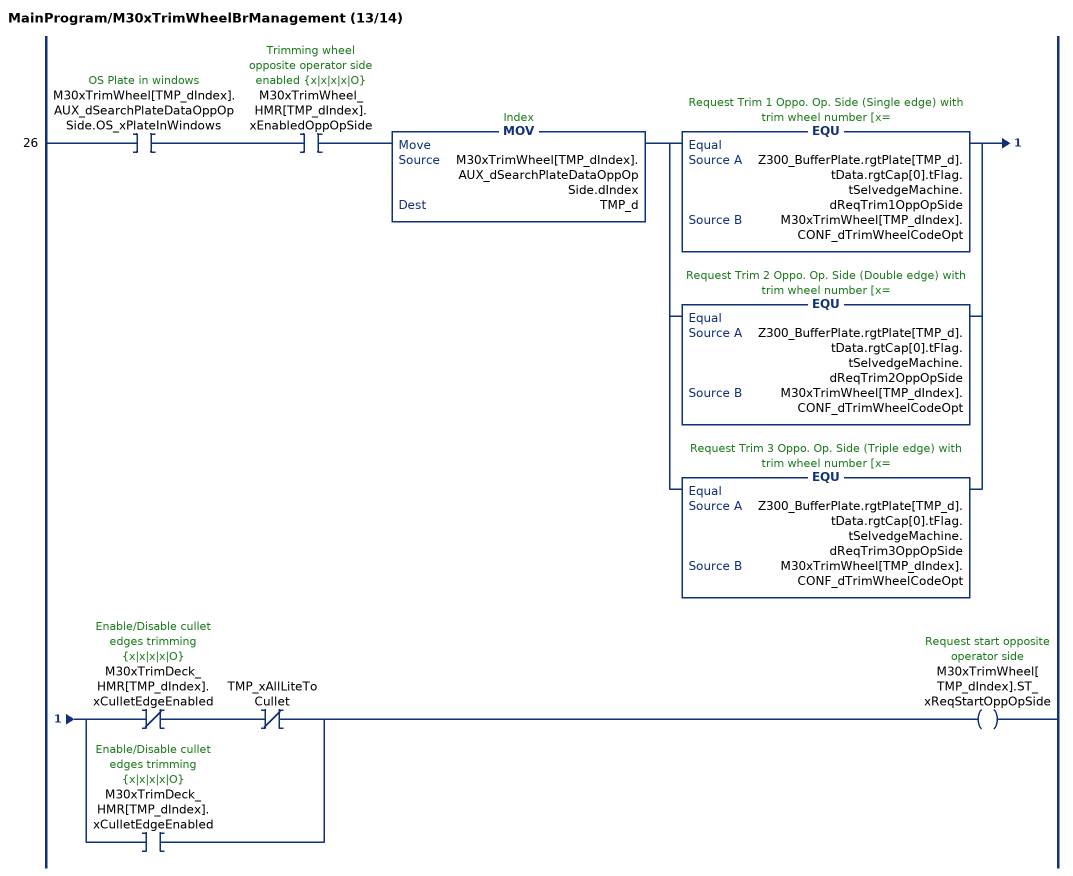
   26: XIC(M30xTrimWheel[TMP_dIndex].AUX_dSearchPlateDataOppOpSide.OS_xPlateInWindows)XIC(M30xTrimWheel_HMR[TMP_dIndex].xEnabledOppOpSide)MOV(M30xTrimWheel[TMP_dIndex].AUX_dSearchPlateDataOppOpSide.dIndex,TMP_d)[EQU(Z300_BufferPlate.rgtPlate[TMP_d].tData.rgtCap[0].tFlag.tSelvedgeMachine.dReqTrim1OppOpSide,M30xTrimWheel[TMP_dIndex].CONF_dTrimWheelCodeOpt) ,EQU(Z300_BufferPlate.rgtPlate[TMP_d].tData.rgtCap[0].tFlag.tSelvedgeMachine.dReqTrim2OppOpSide,M30xTrimWheel[TMP_dIndex].CONF_dTrimWheelCodeOpt) ,EQU(Z300_BufferPlate.rgtPlate[TMP_d].tData.rgtCap[0].tFlag.tSelvedgeMachine.dReqTrim3OppOpSide,M30xTrimWheel[TMP_dIndex].CONF_dTrimWheelCodeOpt) ][XIO(M30xTrimDeck_HMR[TMP_dIndex].xCulletEdgeEnabled) XIO(TMP_xAllLiteToCullet) ,XIC(M30xTrimDeck_HMR[TMP_dIndex].xCulletEdgeEnabled) ]OTE(M30xTrimWheel[TMP_dIndex].ST_xReqStartOppOpSide);
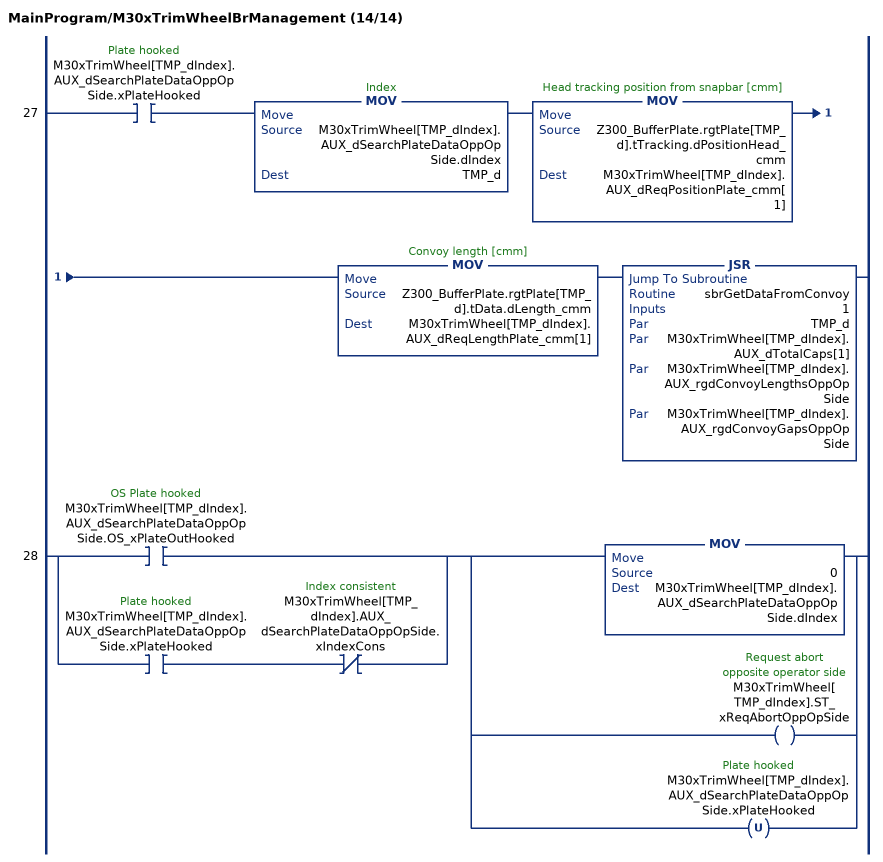
   27: XIC(M30xTrimWheel[TMP_dIndex].AUX_dSearchPlateDataOppOpSide.xPlateHooked)MOV(M30xTrimWheel[TMP_dIndex].AUX_dSearchPlateDataOppOpSide.dIndex,TMP_d)MOV(Z300_BufferPlate.rgtPlate[TMP_d].tTracking.dPositionHead_cmm,M30xTrimWheel[TMP_dIndex].AUX_dReqPositionPlate_cmm[1])MOV(Z300_BufferPlate.rgtPlate[TMP_d].tData.dLength_cmm,M30xTrimWheel[TMP_dIndex].AUX_dReqLengthPlate_cmm[1])JSR(sbrGetDataFromConvoy,1,TMP_d,M30xTrimWheel[TMP_dIndex].AUX_dTotalCaps[1],M30xTrimWheel[TMP_dIndex].AUX_rgdConvoyLengthsOppOpSide,M30xTrimWheel[TMP_dIndex].AUX_rgdConvoyGapsOppOpSide);
   28: [XIC(M30xTrimWheel[TMP_dIndex].AUX_dSearchPlateDataOppOpSide.OS_xPlateOutHooked) ,XIC(M30xTrimWheel[TMP_dIndex].AUX_dSearchPlateDataOppOpSide.xPlateHooked) XIO(M30xTrimWheel[TMP_dIndex].AUX_dSearchPlateDataOppOpSide.xIndexCons) ][MOV(0,M30xTrimWheel[TMP_dIndex].AUX_dSearchPlateDataOppOpSide.dIndex) ,OTE(M30xTrimWheel[TMP_dIndex].ST_xReqAbortOppOpSide) ,OTU(M30xTrimWheel[TMP_dIndex].AUX_dSearchPlateDataOppOpSide.xPlateHooked) ];
END_ROUTINE

ROUTINE M30xTrimWheelTrManagement   (* ladder *)
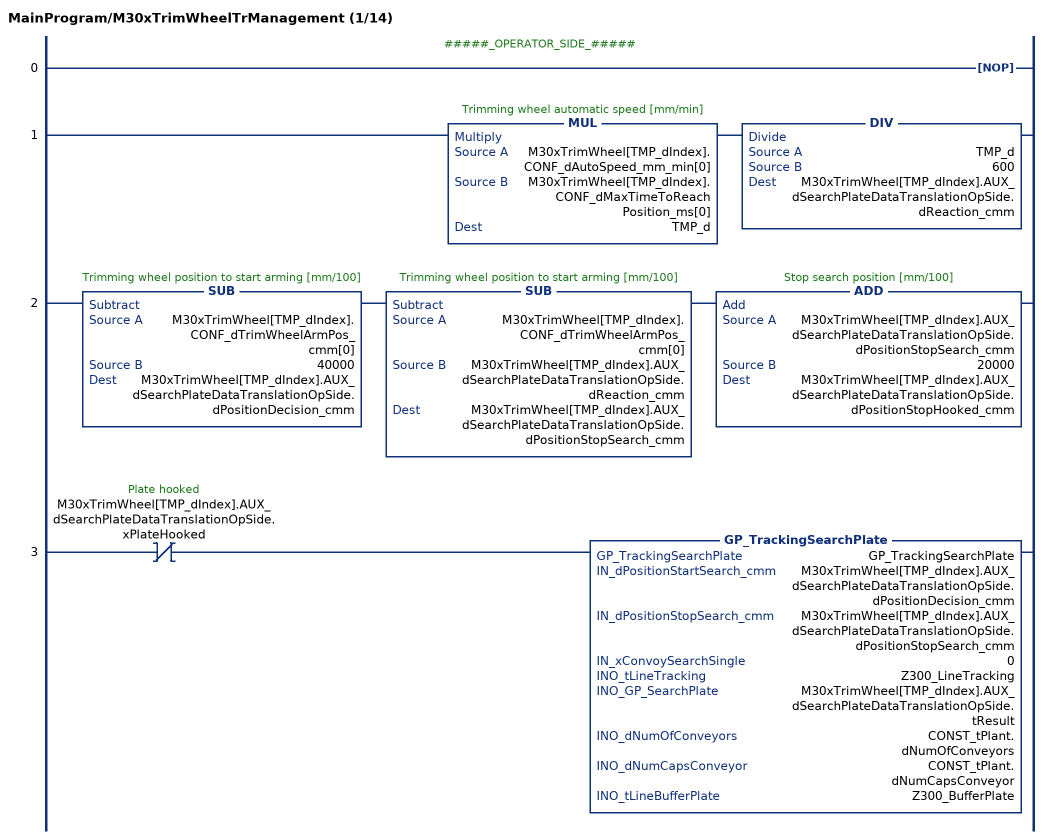
   // #####_OPERATOR_SIDE_#####
   0: NOP();
   1: MUL(M30xTrimWheel[TMP_dIndex].CONF_dAutoSpeed_mm_min[0],M30xTrimWheel[TMP_dIndex].CONF_dMaxTimeToReachPosition_ms[0],TMP_d)DIV(TMP_d,600,M30xTrimWheel[TMP_dIndex].AUX_dSearchPlateDataTranslationOpSide.dReaction_cmm);
   2: SUB(M30xTrimWheel[TMP_dIndex].CONF_dTrimWheelArmPos_cmm[0],40000,M30xTrimWheel[TMP_dIndex].AUX_dSearchPlateDataTranslationOpSide.dPositionDecision_cmm)SUB(M30xTrimWheel[TMP_dIndex].CONF_dTrimWheelArmPos_cmm[0],M30xTrimWheel[TMP_dIndex].AUX_dSearchPlateDataTranslationOpSide.dReaction_cmm,M30xTrimWheel[TMP_dIndex].AUX_dSearchPlateDataTranslationOpSide.dPositionStopSearch_cmm)ADD(M30xTrimWheel[TMP_dIndex].AUX_dSearchPlateDataTranslationOpSide.dPositionStopSearch_cmm,20000,M30xTrimWheel[TMP_dIndex].AUX_dSearchPlateDataTranslationOpSide.dPositionStopHooked_cmm);
   3: XIO(M30xTrimWheel[TMP_dIndex].AUX_dSearchPlateDataTranslationOpSide.xPlateHooked)GP_TrackingSearchPlate(GP_TrackingSearchPlate,M30xTrimWheel[TMP_dIndex].AUX_dSearchPlateDataTranslationOpSide.dPositionDecision_cmm,M30xTrimWheel[TMP_dIndex].AUX_dSearchPlateDataTranslationOpSide.dPositionStopSearch_cmm,0,Z300_LineTracking,M30xTrimWheel[TMP_dIndex].AUX_dSearchPlateDataTranslationOpSide.tResult,CONST_tPlant.dNumOfConveyors,CONST_tPlant.dNumCapsConveyor,Z300_BufferPlate);
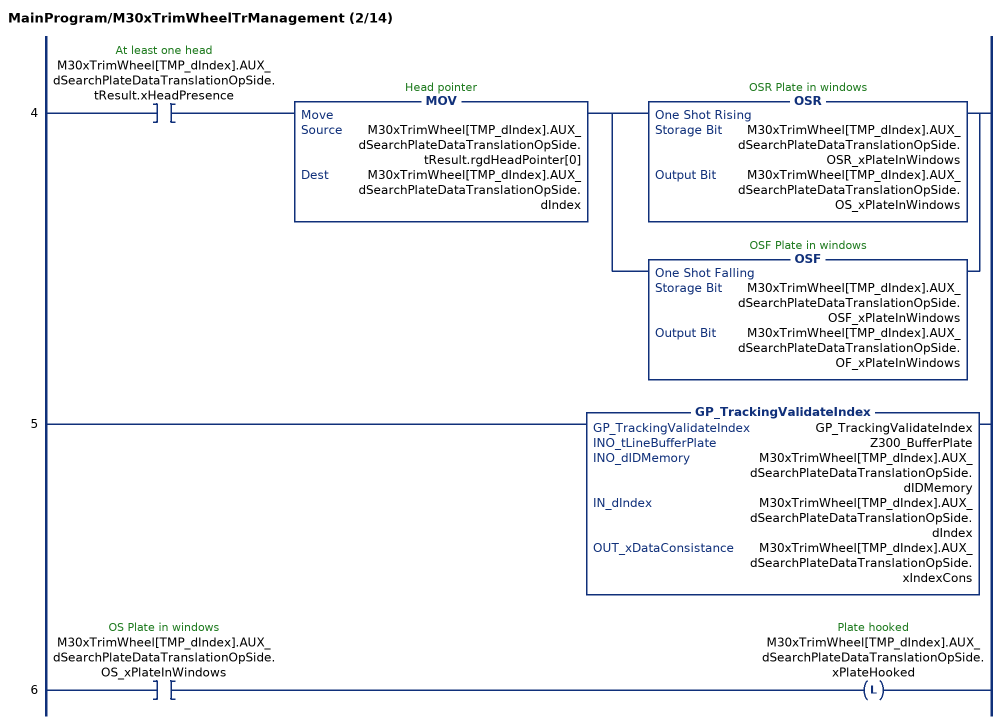
   4: XIC(M30xTrimWheel[TMP_dIndex].AUX_dSearchPlateDataTranslationOpSide.tResult.xHeadPresence)MOV(M30xTrimWheel[TMP_dIndex].AUX_dSearchPlateDataTranslationOpSide.tResult.rgdHeadPointer[0],M30xTrimWheel[TMP_dIndex].AUX_dSearchPlateDataTranslationOpSide.dIndex)[OSR(M30xTrimWheel[TMP_dIndex].AUX_dSearchPlateDataTranslationOpSide.OSR_xPlateInWindows,M30xTrimWheel[TMP_dIndex].AUX_dSearchPlateDataTranslationOpSide.OS_xPlateInWindows) ,OSF(M30xTrimWheel[TMP_dIndex].AUX_dSearchPlateDataTranslationOpSide.OSF_xPlateInWindows,M30xTrimWheel[TMP_dIndex].AUX_dSearchPlateDataTranslationOpSide.OF_xPlateInWindows) ];
   5: GP_TrackingValidateIndex(GP_TrackingValidateIndex,Z300_BufferPlate,M30xTrimWheel[TMP_dIndex].AUX_dSearchPlateDataTranslationOpSide.dIDMemory,M30xTrimWheel[TMP_dIndex].AUX_dSearchPlateDataTranslationOpSide.dIndex,M30xTrimWheel[TMP_dIndex].AUX_dSearchPlateDataTranslationOpSide.xIndexCons);
   6: XIC(M30xTrimWheel[TMP_dIndex].AUX_dSearchPlateDataTranslationOpSide.OS_xPlateInWindows)OTL(M30xTrimWheel[TMP_dIndex].AUX_dSearchPlateDataTranslationOpSide.xPlateHooked);
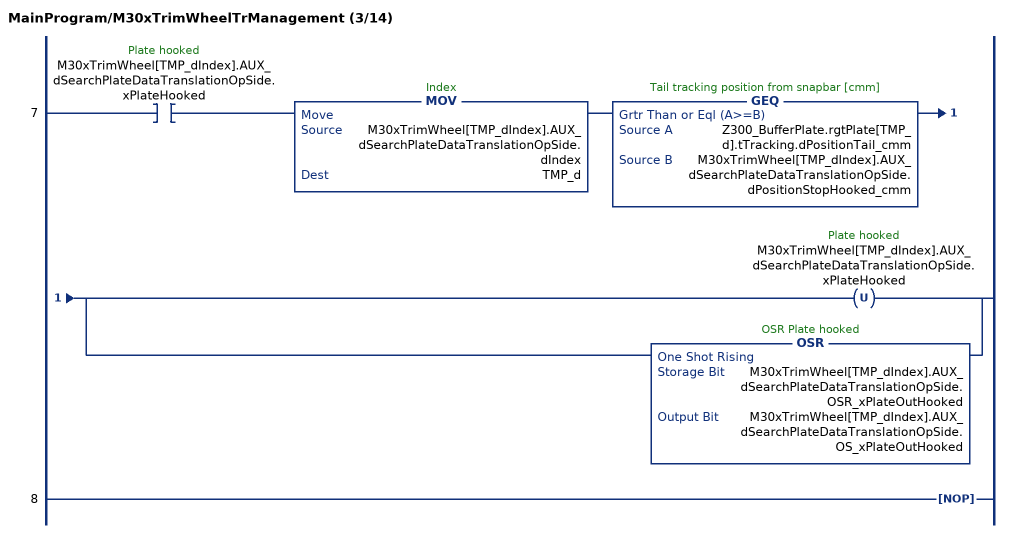
   7: XIC(M30xTrimWheel[TMP_dIndex].AUX_dSearchPlateDataTranslationOpSide.xPlateHooked)MOV(M30xTrimWheel[TMP_dIndex].AUX_dSearchPlateDataTranslationOpSide.dIndex,TMP_d)GEQ(Z300_BufferPlate.rgtPlate[TMP_d].tTracking.dPositionTail_cmm,M30xTrimWheel[TMP_dIndex].AUX_dSearchPlateDataTranslationOpSide.dPositionStopHooked_cmm)[OTU(M30xTrimWheel[TMP_dIndex].AUX_dSearchPlateDataTranslationOpSide.xPlateHooked) ,OSR(M30xTrimWheel[TMP_dIndex].AUX_dSearchPlateDataTranslationOpSide.OSR_xPlateOutHooked,M30xTrimWheel[TMP_dIndex].AUX_dSearchPlateDataTranslationOpSide.OS_xPlateOutHooked) ];
   8: NOP();
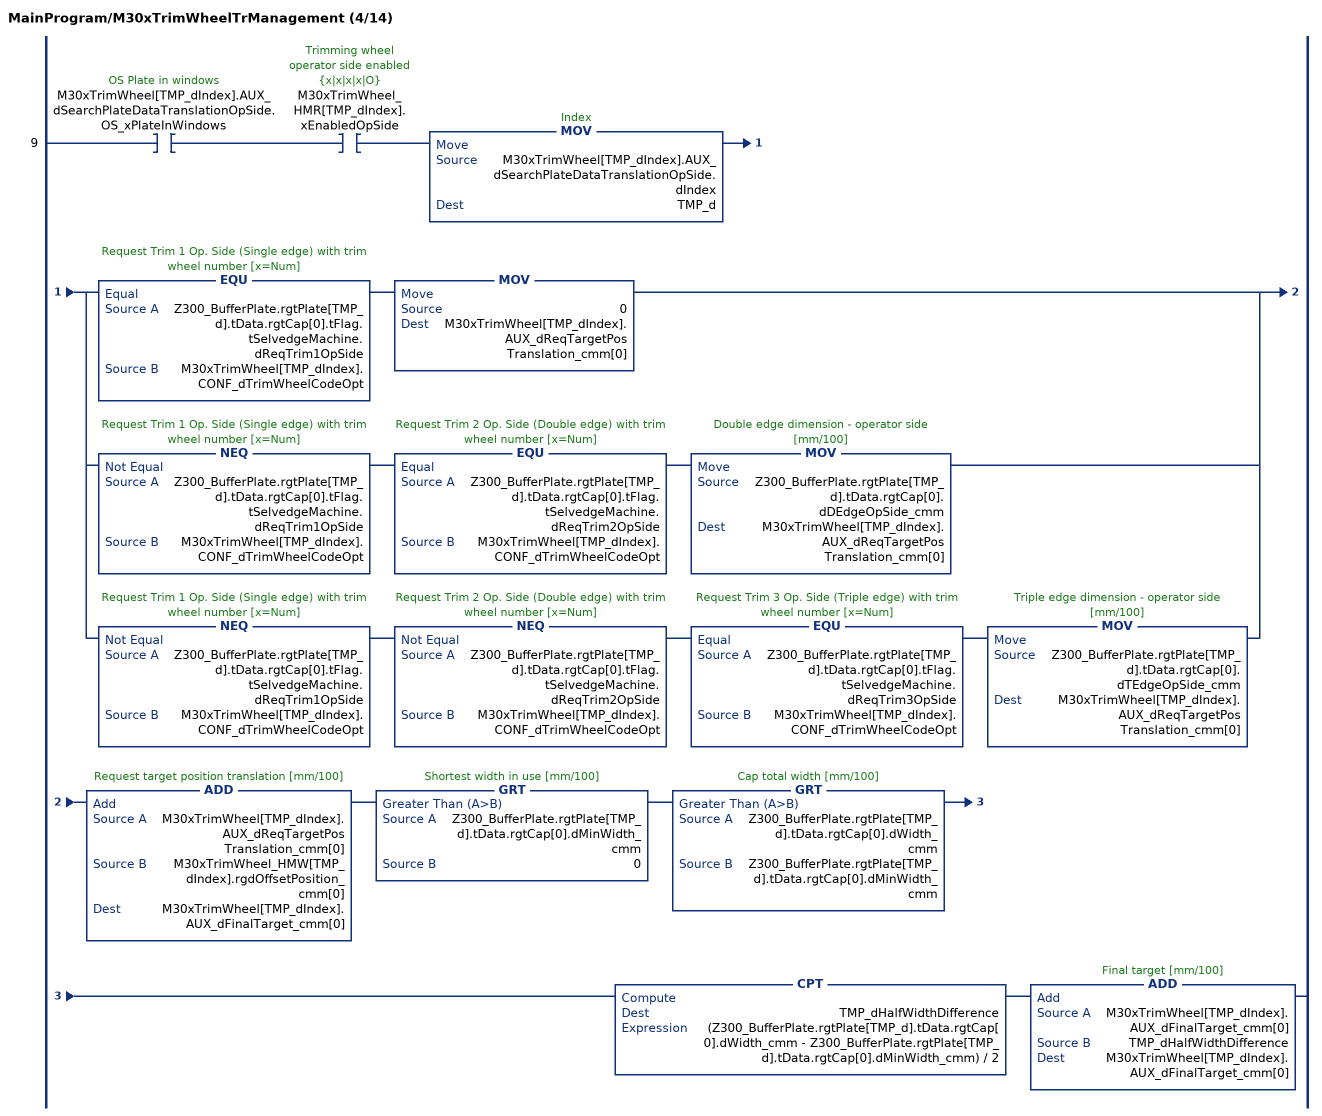
   9: XIC(M30xTrimWheel[TMP_dIndex].AUX_dSearchPlateDataTranslationOpSide.OS_xPlateInWindows)XIC(M30xTrimWheel_HMR[TMP_dIndex].xEnabledOpSide)MOV(M30xTrimWheel[TMP_dIndex].AUX_dSearchPlateDataTranslationOpSide.dIndex,TMP_d)[EQU(Z300_BufferPlate.rgtPlate[TMP_d].tData.rgtCap[0].tFlag.tSelvedgeMachine.dReqTrim1OpSide,M30xTrimWheel[TMP_dIndex].CONF_dTrimWheelCodeOpt) MOV(0,M30xTrimWheel[TMP_dIndex].AUX_dReqTargetPosTranslation_cmm[0]) ,NEQ(Z300_BufferPlate.rgtPlate[TMP_d].tData.rgtCap[0].tFlag.tSelvedgeMachine.dReqTrim1OpSide,M30xTrimWheel[TMP_dIndex].CONF_dTrimWheelCodeOpt) EQU(Z300_BufferPlate.rgtPlate[TMP_d].tData.rgtCap[0].tFlag.tSelvedgeMachine.dReqTrim2OpSide,M30xTrimWheel[TMP_dIndex].CONF_dTrimWheelCodeOpt) MOV(Z300_BufferPlate.rgtPlate[TMP_d].tData.rgtCap[0].dDEdgeOpSide_cmm,M30xTrimWheel[TMP_dIndex].AUX_dReqTargetPosTranslation_cmm[0]) ,NEQ(Z300_BufferPlate.rgtPlate[TMP_d].tData.rgtCap[0].tFlag.tSelvedgeMachine.dReqTrim1OpSide,M30xTrimWheel[TMP_dIndex].CONF_dTrimWheelCodeOpt) NEQ(Z300_BufferPlate.rgtPlate[TMP_d].tData.rgtCap[0].tFlag.tSelvedgeMachine.dReqTrim2OpSide,M30xTrimWheel[TMP_dIndex].CONF_dTrimWheelCodeOpt) EQU(Z300_BufferPlate.rgtPlate[TMP_d].tData.rgtCap[0].tFlag.tSelvedgeMachine.dReqTrim3OpSide,M30xTrimWheel[TMP_dIndex].CONF_dTrimWheelCodeOpt) MOV(Z300_BufferPlate.rgtPlate[TMP_d].tData.rgtCap[0].dTEdgeOpSide_cmm,M30xTrimWheel[TMP_dIndex].AUX_dReqTargetPosTranslation_cmm[0]) ]ADD(M30xTrimWheel[TMP_dIndex].AUX_dReqTargetPosTranslation_cmm[0],M30xTrimWheel_HMW[TMP_dIndex].rgdOffsetPosition_cmm[0],M30xTrimWheel[TMP_dIndex].AUX_dFinalTarget_cmm[0])GRT(Z300_BufferPlate.rgtPlate[TMP_d].tData.rgtCap[0].dMinWidth_cmm,0)GRT(Z300_BufferPlate.rgtPlate[TMP_d].tData.rgtCap[0].dWidth_cmm,Z300_BufferPlate.rgtPlate[TMP_d].tData.rgtCap[0].dMinWidth_cmm)CPT(TMP_dHalfWidthDifference,(Z300_BufferPlate.rgtPlate[TMP_d].tData.rgtCap[0].dWidth_cmm - Z300_BufferPlate.rgtPlate[TMP_d].tData.rgtCap[0].dMinWidth_cmm) / 2)ADD(M30xTrimWheel[TMP_dIndex].AUX_dFinalTarget_cmm[0],TMP_dHalfWidthDifference,M30xTrimWheel[TMP_dIndex].AUX_dFinalTarget_cmm[0]);
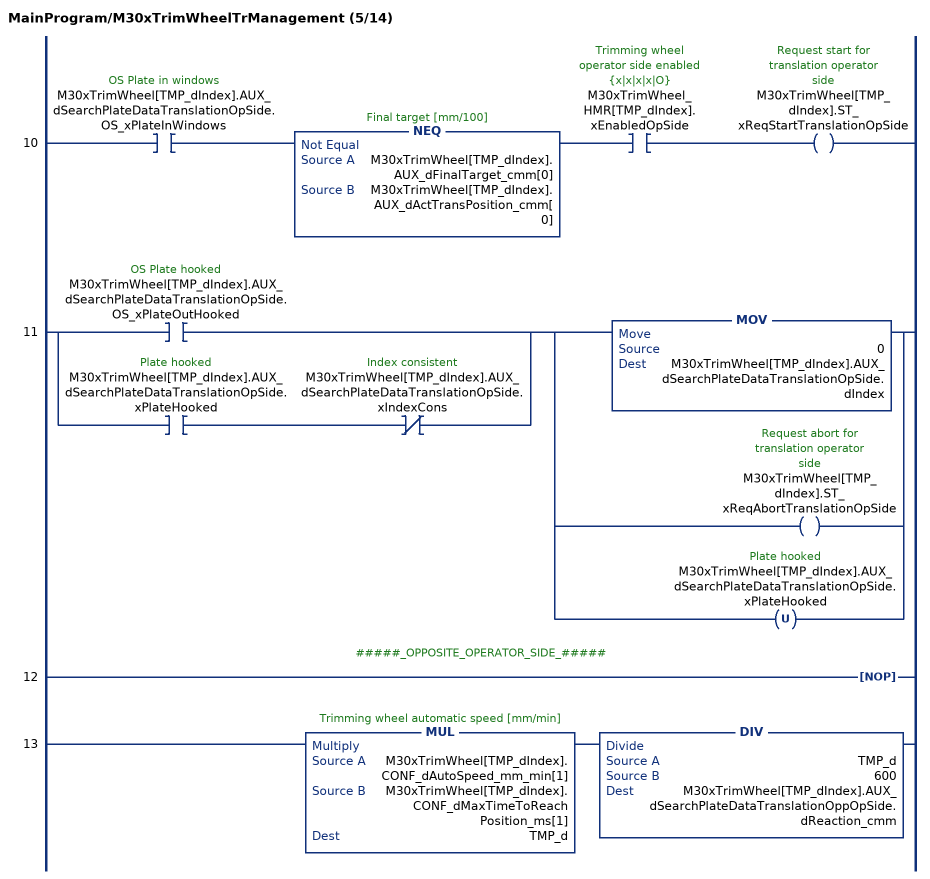
   10: XIC(M30xTrimWheel[TMP_dIndex].AUX_dSearchPlateDataTranslationOpSide.OS_xPlateInWindows)NEQ(M30xTrimWheel[TMP_dIndex].AUX_dFinalTarget_cmm[0],M30xTrimWheel[TMP_dIndex].AUX_dActTransPosition_cmm[0])XIC(M30xTrimWheel_HMR[TMP_dIndex].xEnabledOpSide)OTE(M30xTrimWheel[TMP_dIndex].ST_xReqStartTranslationOpSide);
   11: [XIC(M30xTrimWheel[TMP_dIndex].AUX_dSearchPlateDataTranslationOpSide.OS_xPlateOutHooked) ,XIC(M30xTrimWheel[TMP_dIndex].AUX_dSearchPlateDataTranslationOpSide.xPlateHooked) XIO(M30xTrimWheel[TMP_dIndex].AUX_dSearchPlateDataTranslationOpSide.xIndexCons) ][MOV(0,M30xTrimWheel[TMP_dIndex].AUX_dSearchPlateDataTranslationOpSide.dIndex) ,OTE(M30xTrimWheel[TMP_dIndex].ST_xReqAbortTranslationOpSide) ,OTU(M30xTrimWheel[TMP_dIndex].AUX_dSearchPlateDataTranslationOpSide.xPlateHooked) ];
   // #####_OPPOSITE_OPERATOR_SIDE_#####
   12: NOP();
   13: MUL(M30xTrimWheel[TMP_dIndex].CONF_dAutoSpeed_mm_min[1],M30xTrimWheel[TMP_dIndex].CONF_dMaxTimeToReachPosition_ms[1],TMP_d)DIV(TMP_d,600,M30xTrimWheel[TMP_dIndex].AUX_dSearchPlateDataTranslationOppOpSide.dReaction_cmm);
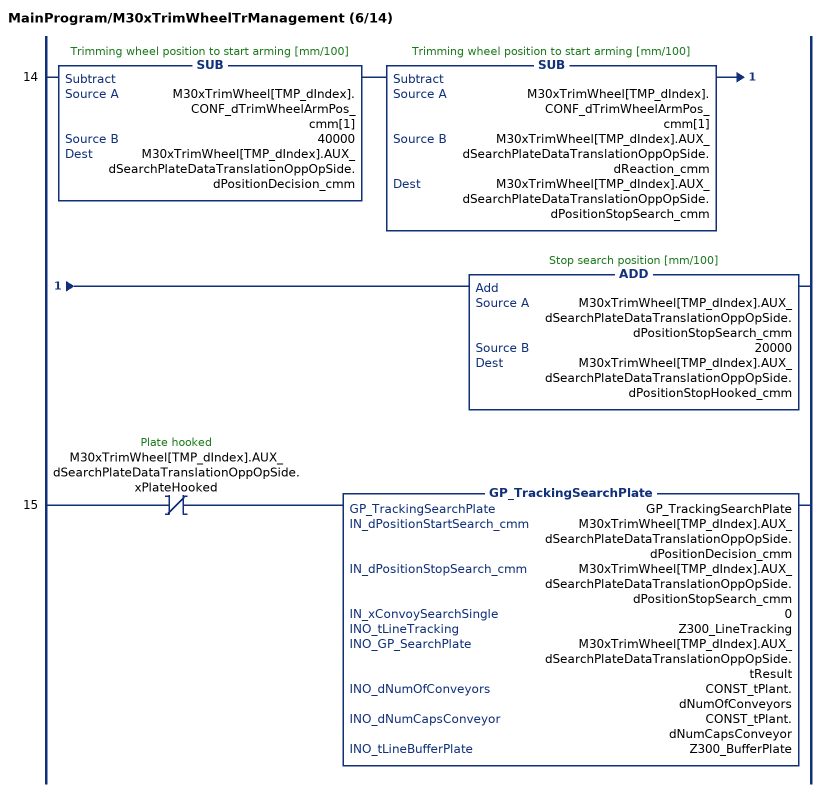
   14: SUB(M30xTrimWheel[TMP_dIndex].CONF_dTrimWheelArmPos_cmm[1],40000,M30xTrimWheel[TMP_dIndex].AUX_dSearchPlateDataTranslationOppOpSide.dPositionDecision_cmm)SUB(M30xTrimWheel[TMP_dIndex].CONF_dTrimWheelArmPos_cmm[1],M30xTrimWheel[TMP_dIndex].AUX_dSearchPlateDataTranslationOppOpSide.dReaction_cmm,M30xTrimWheel[TMP_dIndex].AUX_dSearchPlateDataTranslationOppOpSide.dPositionStopSearch_cmm)ADD(M30xTrimWheel[TMP_dIndex].AUX_dSearchPlateDataTranslationOppOpSide.dPositionStopSearch_cmm,20000,M30xTrimWheel[TMP_dIndex].AUX_dSearchPlateDataTranslationOppOpSide.dPositionStopHooked_cmm);
   15: XIO(M30xTrimWheel[TMP_dIndex].AUX_dSearchPlateDataTranslationOppOpSide.xPlateHooked)GP_TrackingSearchPlate(GP_TrackingSearchPlate,M30xTrimWheel[TMP_dIndex].AUX_dSearchPlateDataTranslationOppOpSide.dPositionDecision_cmm,M30xTrimWheel[TMP_dIndex].AUX_dSearchPlateDataTranslationOppOpSide.dPositionStopSearch_cmm,0,Z300_LineTracking,M30xTrimWheel[TMP_dIndex].AUX_dSearchPlateDataTranslationOppOpSide.tResult,CONST_tPlant.dNumOfConveyors,CONST_tPlant.dNumCapsConveyor,Z300_BufferPlate);
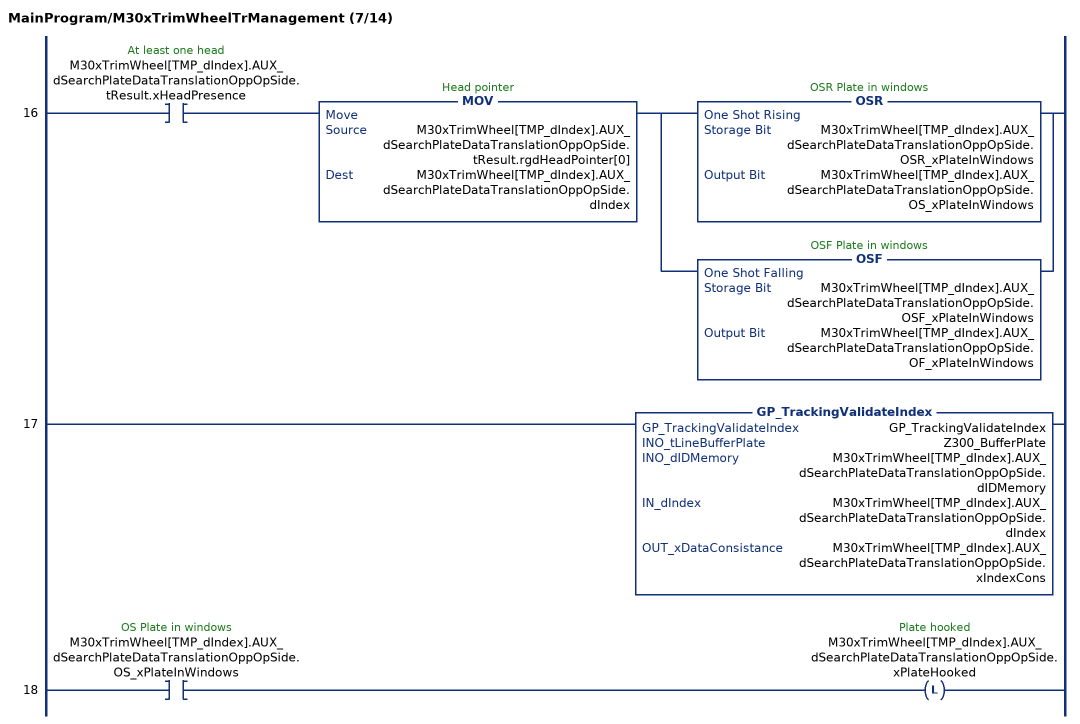
   16: XIC(M30xTrimWheel[TMP_dIndex].AUX_dSearchPlateDataTranslationOppOpSide.tResult.xHeadPresence)MOV(M30xTrimWheel[TMP_dIndex].AUX_dSearchPlateDataTranslationOppOpSide.tResult.rgdHeadPointer[0],M30xTrimWheel[TMP_dIndex].AUX_dSearchPlateDataTranslationOppOpSide.dIndex)[OSR(M30xTrimWheel[TMP_dIndex].AUX_dSearchPlateDataTranslationOppOpSide.OSR_xPlateInWindows,M30xTrimWheel[TMP_dIndex].AUX_dSearchPlateDataTranslationOppOpSide.OS_xPlateInWindows) ,OSF(M30xTrimWheel[TMP_dIndex].AUX_dSearchPlateDataTranslationOppOpSide.OSF_xPlateInWindows,M30xTrimWheel[TMP_dIndex].AUX_dSearchPlateDataTranslationOppOpSide.OF_xPlateInWindows) ];
   17: GP_TrackingValidateIndex(GP_TrackingValidateIndex,Z300_BufferPlate,M30xTrimWheel[TMP_dIndex].AUX_dSearchPlateDataTranslationOppOpSide.dIDMemory,M30xTrimWheel[TMP_dIndex].AUX_dSearchPlateDataTranslationOppOpSide.dIndex,M30xTrimWheel[TMP_dIndex].AUX_dSearchPlateDataTranslationOppOpSide.xIndexCons);
   18: XIC(M30xTrimWheel[TMP_dIndex].AUX_dSearchPlateDataTranslationOppOpSide.OS_xPlateInWindows)OTL(M30xTrimWheel[TMP_dIndex].AUX_dSearchPlateDataTranslationOppOpSide.xPlateHooked);
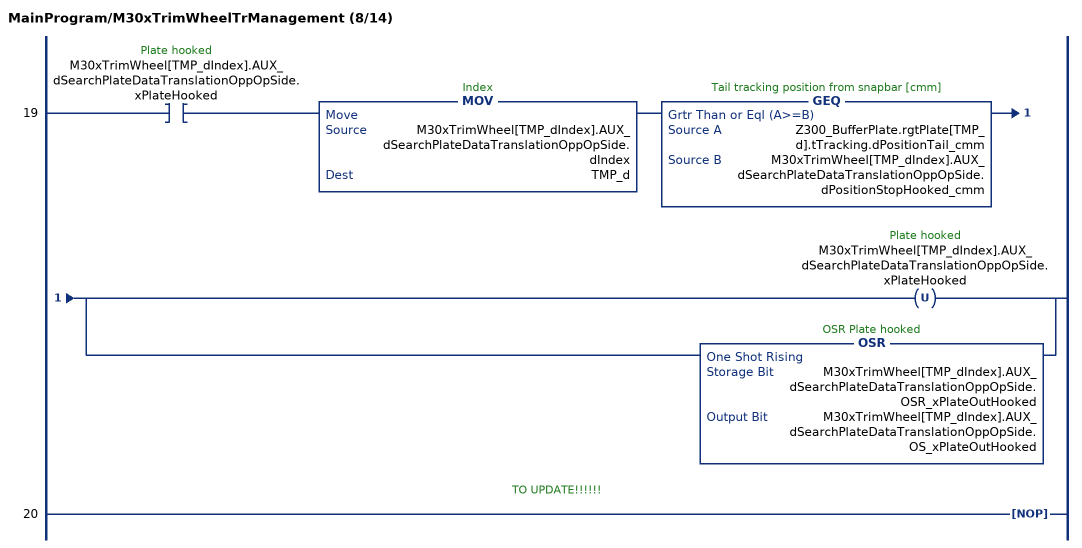
   19: XIC(M30xTrimWheel[TMP_dIndex].AUX_dSearchPlateDataTranslationOppOpSide.xPlateHooked)MOV(M30xTrimWheel[TMP_dIndex].AUX_dSearchPlateDataTranslationOppOpSide.dIndex,TMP_d)GEQ(Z300_BufferPlate.rgtPlate[TMP_d].tTracking.dPositionTail_cmm,M30xTrimWheel[TMP_dIndex].AUX_dSearchPlateDataTranslationOppOpSide.dPositionStopHooked_cmm)[OTU(M30xTrimWheel[TMP_dIndex].AUX_dSearchPlateDataTranslationOppOpSide.xPlateHooked) ,OSR(M30xTrimWheel[TMP_dIndex].AUX_dSearchPlateDataTranslationOppOpSide.OSR_xPlateOutHooked,M30xTrimWheel[TMP_dIndex].AUX_dSearchPlateDataTranslationOppOpSide.OS_xPlateOutHooked) ];
   // TO UPDATE!!!!!!
   20: NOP();
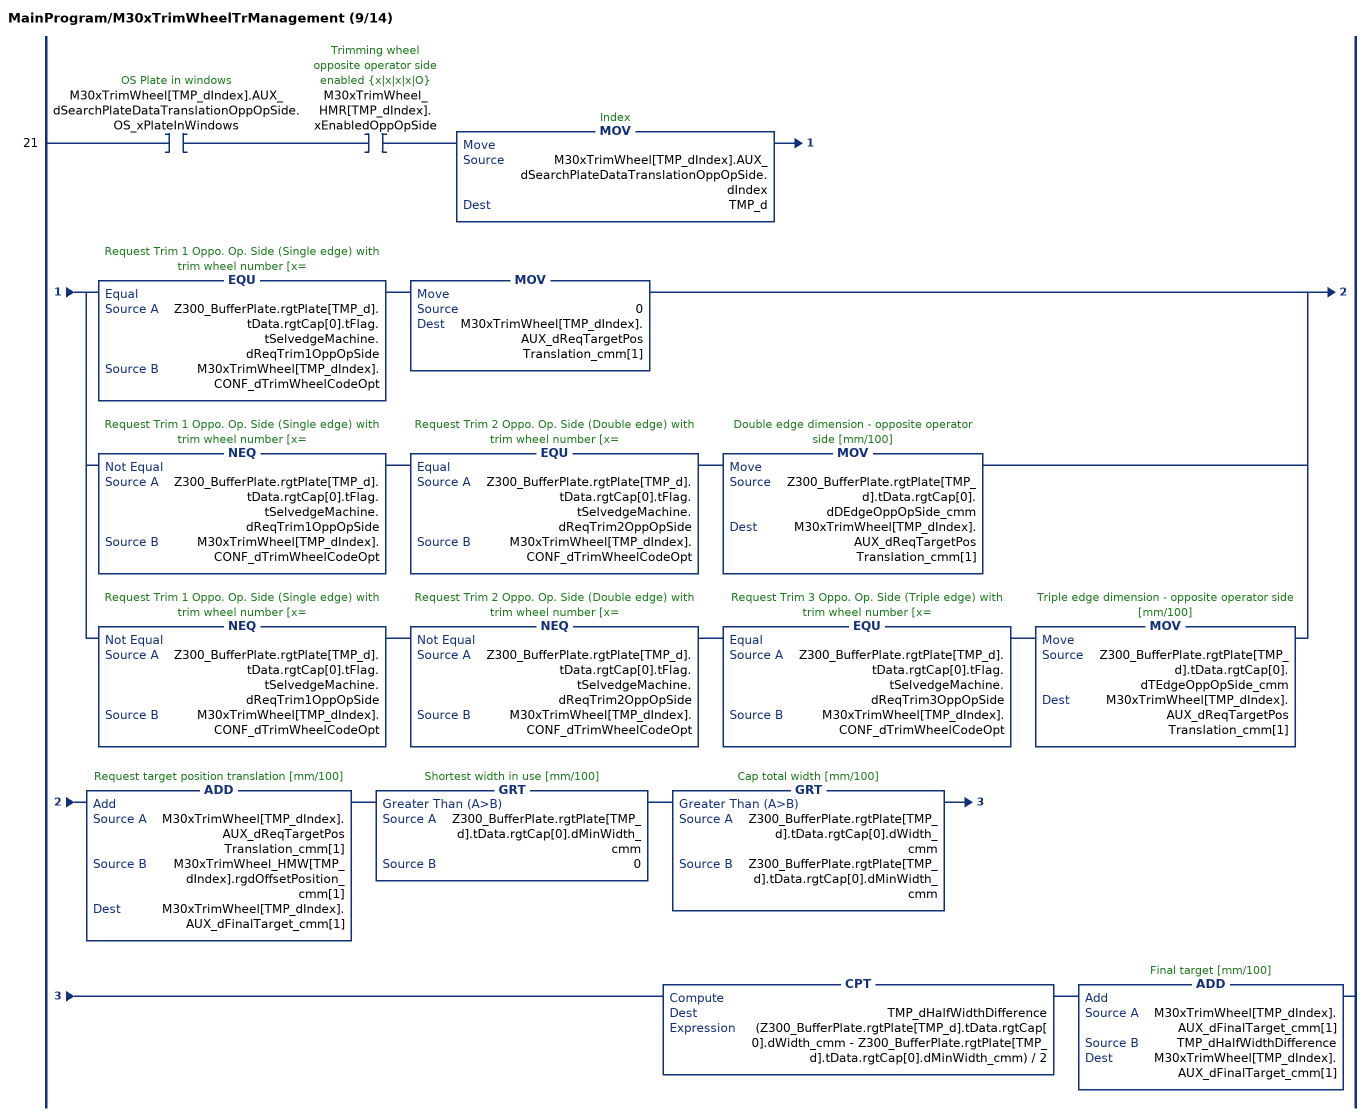
   21: XIC(M30xTrimWheel[TMP_dIndex].AUX_dSearchPlateDataTranslationOppOpSide.OS_xPlateInWindows)XIC(M30xTrimWheel_HMR[TMP_dIndex].xEnabledOppOpSide)MOV(M30xTrimWheel[TMP_dIndex].AUX_dSearchPlateDataTranslationOppOpSide.dIndex,TMP_d)[EQU(Z300_BufferPlate.rgtPlate[TMP_d].tData.rgtCap[0].tFlag.tSelvedgeMachine.dReqTrim1OppOpSide,M30xTrimWheel[TMP_dIndex].CONF_dTrimWheelCodeOpt) MOV(0,M30xTrimWheel[TMP_dIndex].AUX_dReqTargetPosTranslation_cmm[1]) ,NEQ(Z300_BufferPlate.rgtPlate[TMP_d].tData.rgtCap[0].tFlag.tSelvedgeMachine.dReqTrim1OppOpSide,M30xTrimWheel[TMP_dIndex].CONF_dTrimWheelCodeOpt) EQU(Z300_BufferPlate.rgtPlate[TMP_d].tData.rgtCap[0].tFlag.tSelvedgeMachine.dReqTrim2OppOpSide,M30xTrimWheel[TMP_dIndex].CONF_dTrimWheelCodeOpt) MOV(Z300_BufferPlate.rgtPlate[TMP_d].tData.rgtCap[0].dDEdgeOppOpSide_cmm,M30xTrimWheel[TMP_dIndex].AUX_dReqTargetPosTranslation_cmm[1]) ,NEQ(Z300_BufferPlate.rgtPlate[TMP_d].tData.rgtCap[0].tFlag.tSelvedgeMachine.dReqTrim1OppOpSide,M30xTrimWheel[TMP_dIndex].CONF_dTrimWheelCodeOpt) NEQ(Z300_BufferPlate.rgtPlate[TMP_d].tData.rgtCap[0].tFlag.tSelvedgeMachine.dReqTrim2OppOpSide,M30xTrimWheel[TMP_dIndex].CONF_dTrimWheelCodeOpt) EQU(Z300_BufferPlate.rgtPlate[TMP_d].tData.rgtCap[0].tFlag.tSelvedgeMachine.dReqTrim3OppOpSide,M30xTrimWheel[TMP_dIndex].CONF_dTrimWheelCodeOpt) MOV(Z300_BufferPlate.rgtPlate[TMP_d].tData.rgtCap[0].dTEdgeOppOpSide_cmm,M30xTrimWheel[TMP_dIndex].AUX_dReqTargetPosTranslation_cmm[1]) ]ADD(M30xTrimWheel[TMP_dIndex].AUX_dReqTargetPosTranslation_cmm[1],M30xTrimWheel_HMW[TMP_dIndex].rgdOffsetPosition_cmm[1],M30xTrimWheel[TMP_dIndex].AUX_dFinalTarget_cmm[1])GRT(Z300_BufferPlate.rgtPlate[TMP_d].tData.rgtCap[0].dMinWidth_cmm,0)GRT(Z300_BufferPlate.rgtPlate[TMP_d].tData.rgtCap[0].dWidth_cmm,Z300_BufferPlate.rgtPlate[TMP_d].tData.rgtCap[0].dMinWidth_cmm)CPT(TMP_dHalfWidthDifference,(Z300_BufferPlate.rgtPlate[TMP_d].tData.rgtCap[0].dWidth_cmm - Z300_BufferPlate.rgtPlate[TMP_d].tData.rgtCap[0].dMinWidth_cmm) / 2)ADD(M30xTrimWheel[TMP_dIndex].AUX_dFinalTarget_cmm[1],TMP_dHalfWidthDifference,M30xTrimWheel[TMP_dIndex].AUX_dFinalTarget_cmm[1]);
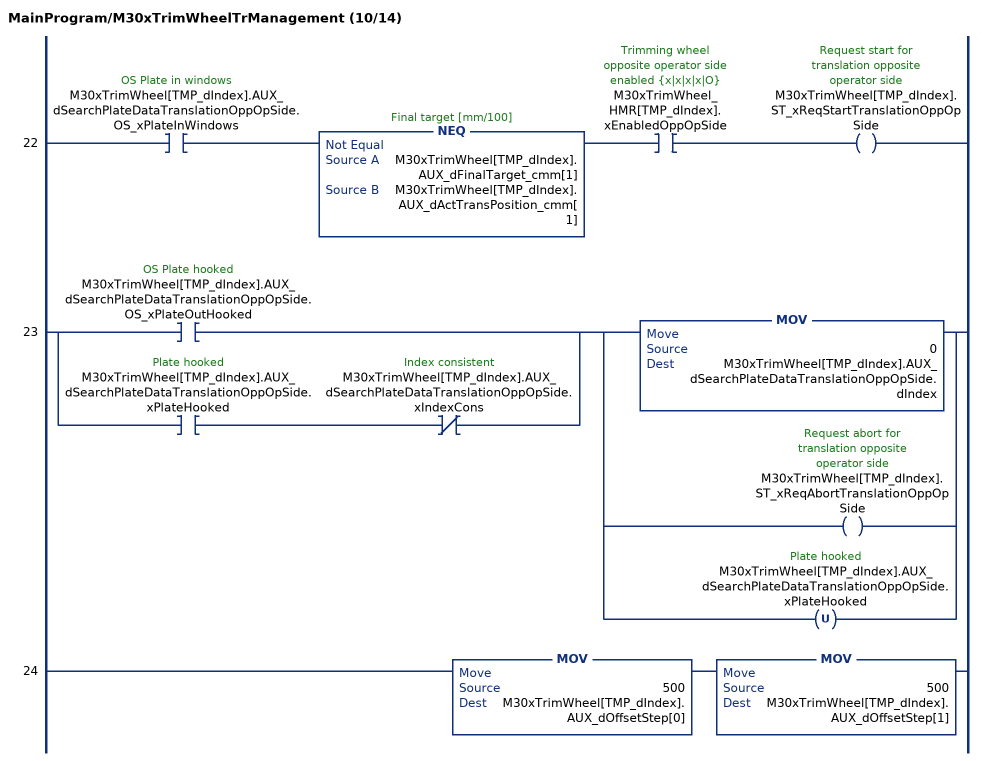
   22: XIC(M30xTrimWheel[TMP_dIndex].AUX_dSearchPlateDataTranslationOppOpSide.OS_xPlateInWindows)NEQ(M30xTrimWheel[TMP_dIndex].AUX_dFinalTarget_cmm[1],M30xTrimWheel[TMP_dIndex].AUX_dActTransPosition_cmm[1])XIC(M30xTrimWheel_HMR[TMP_dIndex].xEnabledOppOpSide)OTE(M30xTrimWheel[TMP_dIndex].ST_xReqStartTranslationOppOpSide);
   23: [XIC(M30xTrimWheel[TMP_dIndex].AUX_dSearchPlateDataTranslationOppOpSide.OS_xPlateOutHooked) ,XIC(M30xTrimWheel[TMP_dIndex].AUX_dSearchPlateDataTranslationOppOpSide.xPlateHooked) XIO(M30xTrimWheel[TMP_dIndex].AUX_dSearchPlateDataTranslationOppOpSide.xIndexCons) ][MOV(0,M30xTrimWheel[TMP_dIndex].AUX_dSearchPlateDataTranslationOppOpSide.dIndex) ,OTE(M30xTrimWheel[TMP_dIndex].ST_xReqAbortTranslationOppOpSide) ,OTU(M30xTrimWheel[TMP_dIndex].AUX_dSearchPlateDataTranslationOppOpSide.xPlateHooked) ];
   24: MOV(500,M30xTrimWheel[TMP_dIndex].AUX_dOffsetStep[0])MOV(500,M30xTrimWheel[TMP_dIndex].AUX_dOffsetStep[1]);
